screen "Inert Gas Conditioning Plant" 1280x800, template "Template_lite"
   on GenerateScreen: "TitleUpdater"()
   GraphicView "Graphic view_20" at 359,634 size 43x62; Picture "Graphic_72"
   GraphicView "Graphic view_52" at 746,80 size 58x108; Picture "Graphic_72"
   GraphicView "Graphic view_63" at 991,218 size 58x108; Picture "Graphic_72"
   GraphicView "Graphic view_64" at 1096,218 size 58x108; Picture "Graphic_72"
   TextField "Text field_64" at 497,462 size 54x22; Text '- OK -'
      Visibility <- "10_DI_DATA_LS_303_LO"
   GraphicView "Graphic view_76" at 53,433 size 168x182; Picture "Graphic_251"
   GraphicView "Graphic view_102" at 12,304 size 58x63; Picture "Graphic_162"
   GraphicView "Graphic view_13" at 724,163 size 182x22; Picture "Graphic_151"
   Group "Group" at 746,80 size 58x108; Picture "Graphic_72"
   GraphicIOField "Graphic I/O field_3" at 188,659 size 60x65; PictureList "Pump Ani"
      ProcessValue <- "10_DI_DATA_P_304_ENBLD"
   GraphicView "Graphic view_18" at 240,683 size 253x11; Picture "Graphic_156"
   GraphicView "Graphic view_89" at 303,257 size 10x13; Picture "Graphic_147"
   GraphicView "Graphic view_59" at 962,301 size 302x22; Picture "Graphic_151"
   GraphicView "Graphic view_5" at 827,163 size 102x22; Picture "Graphic_151"
   Group "Group_2" at 991,218 size 58x108; Picture "Graphic_72"
   TextField "Text field_45" at 989,239 size 60x22; Text 'Closed'
      Visibility <- "10_DI_DATA_CV407_CLSD"
   GraphicView "Graphic view_69" at 124,683 size 68x11; Picture "Graphic_156"
   GraphicView "Graphic view_85" at 235,296 size 33x35; Picture "Graphic_178"
   GraphicView "Graphic view_1" at 259,128 size 301x502; Picture "Graphic_150"
   GraphicView "Graphic view_6" at 870,257 size 18x22; Picture "Graphic_154"
   GraphicView "Graphic view_9" at 689,257 size 188x11; Picture "Graphic_156"
   GraphicView "Graphic view_11" at 424,625 size 12x91; Picture "Graphic_152"
   GraphicView "Graphic view_10" at 424,628 size 19x28; Picture "Graphic_157"
   GraphicView "Graphic view_12" at 440,636 size 106x11; Picture "Graphic_156"
   GraphicView "Graphic view_14" at 817,752 size 20x21; Picture "Graphic_159"
   GraphicView "Graphic view_16" at 635,761 size 188x13; Picture "Graphic_151"
   GraphicIOField "Graphic I/O field_1" at 573,615 size 60x65; PictureList "Pump Ani"
      ProcessValue <- "10_DI_DATA_P_303_ENBLD"
   GraphicView "Graphic view_19" at 471,636 size 106x11; Picture "Graphic_156"
   TextField "Text field_3" at 356,693 size 50x16; Text 'CV-358'
   Group "Group_1" at 359,634 size 43x62; Picture "Graphic_72"
   TextField "Text field_15" at 350,634 size 60x22; Text 'Closed'
      Visibility <- "10_DI_DATA_CV358_CLSD"
   TextField "Text field_16" at 90,573 size 90x22; Text 'PGC Running'
      Visibility <- "10_DI_DATA_E_400_RUN"
   GraphicView "Graphic view_21" at 486,674 size 17x18; Picture "Graphic_153"
   GraphicView "Graphic view_22" at 494,642 size 10x41; Picture "Graphic_152"
   GraphicView "Graphic view_23" at 490,637 size 17x15; Picture "Graphic_161"
   GraphicView "Graphic view_24" at 630,636 size 87x11; Picture "Graphic_156"
   GraphicView "Graphic view_30" at 421,704 size 39x47; Picture "Graphic_162"
   GraphicView "Graphic view_26" at 424,662 size 12x54; Picture "Graphic_152"
   TextField "Text field_1" at 460,713 size 60x22; Text 'Closed'
      Visibility <- "10_DI_DATA_CV341_CLSD"
   TextField "Text field_2" at 460,713 size 60x22; Text 'Opened'
      Visibility <- "10_DI_DATA_CV341_OPN"
   GraphicView "Graphic view_33" at 668,469 size 24x18; Picture "Graphic_155"
   GraphicView "Graphic view_34" at 668,508 size 24x18; Picture "Graphic_166"
   GraphicView "Graphic view_35" at 679,517 size 62x11; Picture "Graphic_156"
   GraphicView "Graphic view_36" at 668,486 size 12x30; Picture "Graphic_152"
   GraphicView "Graphic view_37" at 687,468 size 62x11; Picture "Graphic_156"
   GraphicView "Graphic view_38" at 741,468 size 106x11; Picture "Graphic_156"
   GraphicView "Graphic view_39" at 487,257 size 103x11; Picture "Graphic_156"
   GraphicView "Graphic view_40" at 422,102 size 140x11; Picture "Graphic_156"
   GraphicView "Graphic view_41" at 302,103 size 24x18; Picture "Graphic_155"
   GraphicView "Graphic view_43" at 558,103 size 19x18; Picture "Graphic_154"
   GraphicView "Graphic view_44" at 302,118 size 12x75; Picture "Graphic_152"
   GraphicView "Graphic view_45" at 302,183 size 12x75; Picture "Graphic_152"
   GraphicView "Graphic view_46" at 871,460 size 17x18; Picture "Graphic_153"
   GraphicView "Graphic view_47" at 879,426 size 10x41; Picture "Graphic_152"
   GraphicView "Graphic view_48" at 771,468 size 106x11; Picture "Graphic_156"
   GraphicView "Graphic view_49" at 879,358 size 10x91; Picture "Graphic_152"
   GraphicView "Graphic view_51" at 879,272 size 10x91; Picture "Graphic_152"
   GraphicView "Graphic view_53" at 574,257 size 126x11; Picture "Graphic_156"
   GraphicView "Graphic view_57" at 319,102 size 140x11; Picture "Graphic_156"
   TextField "Text field_4" at 434,743 size 50x16; Text 'CV-341'
   GraphicView "Graphic view_58" at 1062,188 size 19x119; Picture "Graphic_147"
   GraphicView "Graphic view_60" at 1058,159 size 58x63; Picture "Graphic_162"
   TextField "Text field_6" at 995,322 size 50x16; Text 'CV-407'
   GraphicView "Graphic view_61" at 561,250 size 23x16; Picture "Graphic_168"
   GraphicView "Graphic view_62" at 567,179 size 10x77; Picture "Graphic_152"
   TextField "Text field_8" at 1103,322 size 50x16; Text 'CV-411'
   Group "Group_3" at 1096,218 size 58x108; Picture "Graphic_72"
   GraphicView "Graphic view_65" at 1062,151 size 19x23; Picture "Graphic_147"
   TextField "Text field_9" at 1097,239 size 60x22; Text 'Closed'
      Visibility <- "10_DI_DATA_CV411_CLSD"
   TextField "Text field_10" at 1097,239 size 60x22; Text 'Opened'
      Visibility <- "10_DI_DATA_CV411_OPN"
   TextField "Text field_13" at 1115,180 size 60x22; Text 'Opened'
      Visibility <- "10_DI_DATA_CV409_OPN"
   TextField "Text field_17" at 582,680 size 42x16; Text 'P-303'
   TextField "Text field_5" at 1082,214 size 50x16; Text 'CV-409'
   GraphicView "Graphic view_66" at 508,761 size 188x13; Picture "Graphic_151"
   GraphicView "Graphic view_67" at 375,761 size 188x13; Picture "Graphic_151"
   GraphicView "Graphic view_31" at 424,748 size 12x38; Picture "Graphic_152"
   GraphicView "Graphic view_68" at 118,761 size 285x13; Picture "Graphic_151"
   GraphicView "Graphic view_70" at 826,617 size 12x146; Picture "Graphic_147"
   GraphicView "Graphic view_71" at 818,611 size 19x21; Picture "Graphic_169"
   GraphicView "Graphic view_73" at 14,359 size 19x222; Picture "Graphic_147"
   GraphicView "Graphic view_75" at 696,479 size 76x194; Picture "Graphic_173"
   GraphicView "Graphic view_72" at 760,610 size 68x13; Picture "Graphic_151"
   GraphicView "Graphic view_32" at 847,514 size 19x20; Picture "Graphic_169"
   GraphicView "Graphic view_77" at 759,513 size 97x13; Picture "Graphic_151"
   GraphicView "Graphic view_28" at 855,527 size 12x146; Picture "Graphic_147"
   GraphicView "Graphic view_79" at 855,649 size 12x130; Picture "Graphic_147"
   TextField "Text field_24" at 610,79 size 50x16; Text 'CV-405'
   TextField "Text field_27" at 820,266 size 48x16; Text 'FS-350'
   GraphicView "Graphic view_15" at 834,232 size 20x26; Picture "Graphic_79"
   TextField "Text field_40" at 813,209 size 70x22; Text 'No Flow'
      Visibility <- "10_DI_DATA_FS_350_FLW_OK"
   TextField "Text field_41" at 813,209 size 70x22; Text '- Flow -'
      Visibility <- "10_DI_DATA_FS_350_FLW_OK"
   GraphicView "Graphic view_8" at 558,596 size 10x11; Picture "Graphic_159"
   GraphicView "Graphic view_17" at 563,440 size 5x162; Picture "Graphic_147"
   GraphicView "Graphic view_25" at 558,275 size 10x11; Picture "Graphic_169"
   GraphicView "Graphic view_27" at 563,280 size 5x177; Picture "Graphic_147"
   GraphicView "Graphic view_29" at 486,602 size 78x5; Picture "Graphic_151"
   GraphicView "Graphic view_80" at 488,275 size 76x5; Picture "Graphic_151"
   IOField "I/O field_2" at 524,401 size 82x35; FormatPattern 999.9; Unit  %
      ProcessValue <- "12_AI_Data_LIT_304_SCALED"
   TextField "Text field_29" at 669,184 size 56x16; Text 'PIT-416'
   GraphicView "Graphic view_81" at 687,140 size 20x26; Picture "Graphic_36"
   TextField "Text field_25" at 752,442 size 56x16; Text 'TIT-408'
   TextField "Text field_30" at 512,199 size 56x16; Text 'TIT-406'
   GraphicView "Graphic view_82" at 530,137 size 20x26; Picture "Graphic_36"
   TextField "Text field_26" at 824,348 size 56x16; Text 'PIT-353'
   GraphicView "Graphic view_84" at 15,559 size 33x36; Picture "Graphic_177"
   TextField "Text field_7" at 750,184 size 50x16; Text 'CV-406'
   Bar "Bar_1" at 377,282 size 109x327; Unit  %; MinimumValue 0; MaximumValue 100
      ProcessValue <- "12_AI_Data_LIT_304_SCALED"
   TextField "Text field_48" at 16,624 size 112x20; Text 'PG Compressor'
      Appearance <- "10_DI_DATA_E_400_NOK"
   TextField "Text field_34" at 615,534 size 79x34; Text 'Heat Exchanger'
   TextField "Text field_35" at 551,697 size 100x34; Text 'Recirculation Pump'
   TextField "Text field_36" at 402,782 size 61x18; Text 'To Bilge'
   TextField "Text field_37" at 814,782 size 100x18; Text 'To Overboard'
   Group "Group_5" at 396,264 size 74x42
   GraphicView "Graphic view_3" at 429,258 size 15x16; Picture "Graphic_178"
   GraphicView "Graphic view_88" at 434,257 size 55x11; Picture "Graphic_151"
   TextField "Text field_38" at 571,440 size 55x16; Text 'LIT-304'
   TextField "Text field_39" at 269,693 size 56x16; Text 'PIT-358'
   GraphicView "Graphic view_90" at 287,658 size 20x26; Picture "Graphic_36"
   TextField "Text field_28" at 704,774 size 56x16; Text 'PIT-348'
   GraphicView "Graphic view_83" at 722,736 size 20x26; Picture "Graphic_36"
   TextField "Text field_31" at 778,623 size 48x16; Text 'FS-332'
   GraphicView "Graphic view_91" at 801,585 size 20x26; Picture "Graphic_79"
   TextField "Text field_32" at 779,562 size 70x22; Text 'No Flow'
      Visibility <- "10_DI_DATA_FS_332 FLW_OK"
   TextField "Text field_42" at 779,562 size 70x22; Text '- Flow -'
      Visibility <- "10_DI_DATA_FS_332 FLW_OK"
   TextField "Text field_43" at 197,724 size 42x16; Text 'P-304'
   TextField "Text field_44" at 169,740 size 106x20; Text 'Booster Pump'
   GraphicView "Graphic view_2" at 553,163 size 182x22; Picture "Graphic_151"
   TextField "Text field_11" at 989,239 size 60x22; Text 'Opened'
      Visibility <- "10_DI_DATA_CV407_OPN"
   GraphicView "Graphic view_7" at 251,453 size 24x21; Picture "Graphic_107"
   TextField "Text field_46" at 225,501 size 86x16; Text 'E-400-PT002'
   TextField "Text field_47" at 132,408 size 86x16; Text 'E-400-TT002'
   GraphicView "Graphic view_87" at 234,321 size 19x128; Picture "Graphic_147"
   GraphicView "Graphic view_86" at 220,442 size 33x36; Picture "Graphic_159"
   IOField "I/O field_10" at 683,53 size 57x22; FormatPattern 999
      ProcessValue <- "12_AI_Data_CV_405_SCALED"
   IOField "I/O field_11" at 226,482 size 68x18; FormatPattern 999.9; Unit  Bar
      ProcessValue <- "12_AI_Data_E_400_PT002_SCALED"
   IOField "I/O field_13" at 663,119 size 68x18; FormatPattern 99.99; Unit  Bar
      ProcessValue <- "12_AI_Data_PIT_416_SCALED"
   IOField "I/O field_14" at 787,330 size 68x18; FormatPattern 99.99; Unit  Bar
      ProcessValue <- "12_AI_Data_PIT_353_SCALED"
   IOField "I/O field_15" at 704,426 size 68x18; FormatPattern 99.99; Unit  °C
      ProcessValue <- "12_AI_Data_TIT_408_SCALED"
   IOField "I/O field_16" at 698,717 size 68x18; FormatPattern 99.99; Unit  Bar
      ProcessValue <- "12_AI_Data_PIT_348_SCALED"
   IOField "I/O field_7" at 263,638 size 68x18; FormatPattern 99.99; Unit  Bar
      ProcessValue <- "12_AI_Data_PIT_358_SCALED"
   TextField "Text field_57" at 1021,112 size 90x32; Text 'Vent To Atmosphere'
   TextField "Text field_58" at 608,3 size 150x18; Text 'Vent To Atmosphere'
   IOField "I/O field_1" at 143,392 size 68x18; FormatPattern 999.9; Unit  °C
      ProcessValue <- "12_AI_Data_E_400_TE002_SCALED"
   GraphicView "Graphic view_93" at 491,492 size 24x21; Picture "Graphic_107"
   TextField "Text field_63" at 515,491 size 48x16; Text 'LS-303'
   TextField "Text field_66" at 497,462 size 54x22; Text 'Low Low'
      Visibility <- "10_DI_DATA_LS_303_LO"
   TextField "Text field_90" at 497,462 size 54x22; Text '-LOW-'
      Visibility <- "10_DI_DATA_LS_303_LO"
   GraphicView "Graphic view_94" at 99,304 size 58x63; Picture "Graphic_162"
   TextField "Text field_70" at 125,264 size 60x22; Text 'Opened'
      Visibility <- "10_DI_DATA_CV441_OPN"
   TextField "Text field_71" at 126,288 size 50x16; Text 'CV-441'
   GraphicView "Graphic view_95" at 103,278 size 19x41; Picture "Graphic_147"
   TextField "Text field_72" at 93,222 size 65x32; Text 'Ambient Air Inlet'
   GraphicView "Graphic view_96" at 86,364 size 36x39; Picture "Graphic_159"
   GraphicView "Graphic view_97" at 28,382 size 70x22; Picture "Graphic_151"
   TextField "Text field_69" at 125,264 size 60x22; Text 'Closed'
      Visibility <- "10_DI_DATA_CV441_CLSD"
   TextField "Text field_12" at 1115,180 size 60x22; Text 'Closed'
      Visibility <- "10_DI_DATA_CV409_CLSD"
   GraphicView "Graphic view_98" at 0,278 size 33x35; Picture "Graphic_169"
   GraphicView "Graphic view_99" at 856,330 size 23x20; Picture "Graphic_255"
   GraphicView "Graphic view_100" at 728,443 size 20x26; Picture "Graphic_36"
   TextField "Text field_33" at 744,96 size 60x22; Text 'Closed'
      Visibility <- "10_DI_DATA_CV406_CLSD"
   TextField "Text field_14" at 744,96 size 60x22; Text 'Opened'
      Visibility <- "10_DI_DATA_CV406_OPN"
   TextField "Text field_18" at 950,356 size 149x23; Text 'Hazardous Area'
   GraphicView "Graphic view_4" at 1204,277 size 20x26; Picture "Graphic_36"
   IOField "I/O field_3" at 1180,257 size 68x18; FormatPattern 99.99; Unit  Bar
      ProcessValue <- "20_TANKS_IP_DATA_RIO_06_FIRST_TANK_DECK_IG_PRESS"
   TextField "Text field_20" at 1186,322 size 56x16; Text 'PIT-415'
   GraphicView "Graphic view_50" at 100,253 size 26x26; Picture "Graphic_261"
   GraphicView "Graphic view_74" at 549,146 size 18x54; Picture "Graphic_281"
   GraphicView "Graphic view_78" at 256,278 size 17x59; Picture "Graphic_281"
   GraphicView "Graphic view_101" at 213,397 size 23x20; Picture "Graphic_255"
   TextField "Text field_56" at 1229,342 size 44x32; Text 'To BWTS'
   TextField "Text field_60" at 661,356 size 94x23; Text 'Safe Area'
   IOField "I/O field_4" at 683,37 size 57x22; FormatPattern 999
      ProcessValue <- "16_AQ_Data_CV405_CNTRL"
   TextField "Text field_106" at 752,38 size 59x18; Text 'OPENED'
   GraphicView "Graphic view_103" at 14,298 size 19x22; Picture "Graphic_147"
   TextField "Text field_73" at 34,288 size 50x16; Text 'CV-401'
   TextField "Text field_74" at 30,264 size 60x22; Text 'Opened'
      Visibility <- "10_DI_Data_CV401_OPN"
   TextField "Text field_75" at 30,264 size 60x22; Text 'Closed'
      Visibility <- "10_DI_Data_CV401_CLSD"
   Button "HmiScreenItemData_13" at 4,669 size 121x40; TextOn 'IGG Plant'; TextOff 'Fresh Water System'; Authorization "Operate"
      on Release: ActivateScreen("Fresh Water System", 0)
      Appearance <- "10 DI_DATA_P305_ENBLD"
   Button "HmiScreenItemData_11" at 3,745 size 122x41; TextOn 'IGG Plant'; TextOff 'Cooling System'; Authorization "Operate"
      on Release: ActivateScreen("Cooling System", 0)
   TextField "Text field_22" at 90,573 size 90x22; Text 'PGC Loaded'
      Visibility <- "10_DI_DATA_E_400_RUN"
   Button "HmiScreenItemData_12" at 46,424 size 177x198; TextOn 'IGG Plant'; TextOff 'Text'; Authorization "Operate"
      on Release: ActivateScreen("PGC System", 0)
   TextField "Text field_23" at 350,634 size 60x22; Text 'Opened'
      Visibility <- "10_DI_DATA_CV358_OPN"
   GraphicView "Graphic view_54" at 588,60 size 19x108; Picture "Graphic_147"
   GraphicView "Graphic view_55" at 586,28 size 95x54; Picture "Graphic_167"
   GraphicView "Graphic view_56" at 588,8 size 19x33; Picture "Graphic_147"
   IOField "I/O field_12" at 506,119 size 68x18; FormatPattern 99.99; Unit  °C
      ProcessValue <- "12_AI_Data_TIT_406_SCALED"
   GraphicView "Graphic view_42" at 567,116 size 10x51; Picture "Graphic_152"
   TextField "Text field_76" at 618,40 size 30x22; Text 'A'
      Visibility <- "19_AUTO_CMNDS_Data_CV405_PID_MDLTG"
   GraphicView "Logo" at 1,1 size 219x60; Picture "Logo of IGG HMI"
   Button "HmiScreenItemData_1" at 1,50 size 150x43; TextOn 'Back'; TextOff 'Main Index'
      on Release: ActivateScreen("02 Main Index", 0)
   GraphicView "Graphic view_92" at 925,164 size 33x36; Picture "Graphic_169"
   Button "HmiScreenItemData_2" at 1128,64 size 150x43; TextOn 'Back'; TextOff 'GCU Setup'; Authorization "Operate"
      on Release: ActivateScreen("Inert Gas Conditioning Setup", 0)
   DateTimeField "HmiScreenItemData_17" at 1175,0 size 105x30
   DateTimeField "HmiScreenItemData" at 1175,30 size 105x30
   GraphicView "Graphic view_106" at 939,194 size 19x100; Picture "Graphic_147"
   GraphicView "Graphic view_104" at 940,285 size 33x37; Picture "Graphic_177"
   Button "HmiScreenItemData_9" at 930,410 size 340x30; TextOn 'Back'; TextOff 'GCU CONTROL'
      Visibility <- "150_GCU_LCL_CNTRL_DB_LCL_CNTRL_ACTV"
   Line "Line_2" at 1246,550 size 0x80
      Visibility <- "150_GCU_LCL_CNTRL_DB_LCL_CNTRL_ACTV"
   Line "Line_3" at 1080,630 size 166x0
      Visibility <- "150_GCU_LCL_CNTRL_DB_LCL_CNTRL_ACTV"
   Button "HmiScreenItemData_4" at 930,610 size 150x40; TextOn 'Back'; TextOff 'Stop'; Authorization "Commissioning"
      on Press: function_b14e0dd5("150_GCU_LCL_CNTRL_DB_STOP", 0)
      Visibility <- "150_GCU_LCL_CNTRL_DB_LCL_CNTRL_ACTV"
   Line "Line_7" at 1080,530 size 145x0
      Visibility <- "150_GCU_LCL_CNTRL_DB_LCL_CNTRL_ACTV"
   Circle "Circle_20" at 1225,510 size 40x40
      Visibility <- "150_GCU_LCL_CNTRL_DB_LCL_CNTRL_ACTV"
      Appearance <- "150_GCU_LCL_CNTRL_DB_RUN_WITH_AIR"
   Button "HmiScreenItemData_3" at 930,510 size 150x40; TextOn 'Back'; TextOff 'Start With Air'; Authorization "Commissioning"
      on Press: function_b14e0dd5("150_GCU_LCL_CNTRL_DB_STRT_AIR", 0)
      Visibility <- "150_GCU_LCL_CNTRL_DB_LCL_CNTRL_ACTV"
   Button "HmiScreenItemData_5" at 930,450 size 340x40; TextOn 'Back'; TextOff 'Start'; TextList "GCU_LCL"; Authorization "Commissioning"
      on Press: InvertBit("150_GCU_LCL_CNTRL_DB_LCL_CNTRL_ACTV")
      Visibility <- "150_GCU_LCL_CNTRL_DB_LCL_CNTRL_ACTV"
      ProcessValue <- "150_GCU_LCL_CNTRL_DB_LCL_CNTRL_ACTV"
   Button "HmiScreenItemData_6" at 930,560 size 150x40; TextOn 'Back'; TextOff 'Start With IG'; Authorization "Commissioning"
      on Press: function_b14e0dd5("150_GCU_LCL_CNTRL_DB_STRT_IG", 0)
      Visibility <- "150_GCU_LCL_CNTRL_DB_LCL_CNTRL_ACTV"
   Line "Line_6" at 1080,580 size 145x0
      Visibility <- "150_GCU_LCL_CNTRL_DB_LCL_CNTRL_ACTV"
   Circle "Circle_1" at 1225,560 size 40x40
      Visibility <- "150_GCU_LCL_CNTRL_DB_LCL_CNTRL_ACTV"
      Appearance <- "150_GCU_LCL_CNTRL_DB_RUN_WITH_IG"
   Button "HmiScreenItemData_7" at 930,660 size 240x40; TextOn 'Back'; TextOff 'Start With Air'; TextList "GTT_OPS"; Authorization "Commissioning"
      on Press: InvertBit("150_GCU_LCL_CNTRL_DB_OPN_ACTV_GTT_VLVS")
      Visibility <- "150_GCU_LCL_CNTRL_DB_LCL_CNTRL_ACTV"
      ProcessValue <- "150_GCU_LCL_CNTRL_DB_OPN_ACTV_GTT_VLVS"
   Circle "Circle_2" at 1225,660 size 40x40
      Visibility <- "150_GCU_LCL_CNTRL_DB_LCL_CNTRL_ACTV"
      Appearance <- "150_GCU_LCL_CNTRL_DB_OPN_ACTV_GTT_VLVS"
   Line "Line_14" at 1170,680 size 55x0
      Visibility <- "150_GCU_LCL_CNTRL_DB_LCL_CNTRL_ACTV"
   Group "Group_4" at 187,631 size 60x25
   Group "Group_6" at 573,588 size 60x25
   IOField "I/O field_34" at 664,96 size 66x23; FormatPattern 99.9; Unit  Bar
      ProcessValue <- "19_AUTO_CMNDS_Data_PIT416_CMND_Target"
      Appearance <- "19_AUTO_CMNDS_Data_PIT402_Target"
   Group "Group_7" at 214,1 size 373x50
   GraphicView "Graphic view_105" at 1184,288 size 96x48; Picture "Graphic_235"
   Button "HmiScreenItemData_10" at 1178,277 size 102x71; TextOn 'Back'; TextOff 'Text'
      on Press: ActivateScreen("Balast Water Treatment Plant", 0)
   GraphicView "Graphic view_108" at 2,208 size 95x48; Picture "Left Arow"
   Button "HmiScreenItemData_14" at 1,195 size 106x107; TextOn 'Back'; TextOff 'Text'
      on Press: ActivateScreen("Inert Gas Generator Plant", 0)
   Button "HmiScreenItemData_15" at 1,133 size 158x52; TextOn 'INERT GAS TRANSFER'; TextOff 'Inert Gas Transfer'; TextList "IG Transfer"; Authorization "Operate"
      on Release: ActivateScreen("IG Transfer Mode", 0)
      ProcessValue <- "80_From_HMI_BWT_BYPASS"
   IOField "I/O field_37" at 1070,718 size 79x29; Authorization "Commissioning"; FormatPattern 999; Unit  step
      ProcessValue <- "2110_BTCS_CNTRL_DB_BTCS_STEP"
   Button "HmiScreenItemData_16" at 930,718 size 137x29; TextOn 'Back'; TextOff 'BWTS Step'
   Button "HmiScreenItemData_51" at 930,753 size 137x29; TextOn 'Back'; TextOff 'BWTS State'
   IOField "I/O field_38" at 1070,753 size 79x29; Authorization "Commissioning"; FormatPattern 9; Unit  state
      ProcessValue <- "2110_BTCS_CNTRL_DB_BTCS_STATE"
   Group "Group_9" at 591,11 size 604x305
   Group "Group_12" at 260,515 size 606x260
   Group "Group_13" at 179,634 size 324x58
   GraphicView "Graphic view_107" at 563,347 size 57x58; Picture "Graphic_302"
      Visibility <- "10_DI_DATA_EPB_8S1"
   Group "Group_10" at 389,152 size 96x105
   Group "Group_11" at 239,299 size 243x195
   Group "Group_8" at 384,257 size 504x388
   Button "Button_1" at 655,120 size 84x92; TextOff 'Text'
      on Press: function_efd93a16("PGC Setpoint Protection", 400, 200, -1, -1, 1)
   Button "Button_4" at 578,3 size 84x99; TextOff 'Text'
      on Press: function_efd93a16("CV 405 Grafics", 300, 100, -1, -1, 1)
   Button "HmiScreenItemData_18" at 236,593 size 83x29; TextOn 'Back'; TextOff 'Temp-Trends'
      on Click: function_efd93a16("PGC Temperature Trends", 200, 100, -1, -1, 1)
   Group "Group_14" at 914,406 size 366x378
   Button "Button_3" at 187,631 size 60x25; TextOn 'Alarm'; TextOff 'OK'
      Appearance <- "10_DI_DATA_P_304_OK"
   TextField "Text field_19" at 187,631 size 60x25; Text 'Enabled'
      Visibility <- "14_DQ_DATA_P_304"
      Appearance <- "14_DQ_DATA_P_304"
   Button "Button_2" at 573,588 size 60x25; TextOn 'Alarm'; TextOff 'OK'
      Appearance <- "10_DI_DATA_P_303_OK"
   TextField "Text field_49" at 573,588 size 60x25; Text 'Enabled'
      Visibility <- "14_DQ_DATA_P_303"
      Appearance <- "14_DQ_DATA_P_303"
   Button "HmiScreenItemData_8" at 228,5 size 355x40; TextOn 'Back'; TextOff 'Text'
   TextField "Screen title" at 214,1 size 373x50; Text 'Screen title'
   Circle "Circle_73" at 594,11 size 10x10
      VerticalMovement <- "E-400 Animation_DB_Animation"
      Visibility <- "10_DI_DATA_E_400_RUN"
   Circle "Circle_45" at 592,89 size 10x10
      VerticalMovement <- "E-400 Animation_DB_Animation"
      Visibility <- "10_DI_DATA_E_400_RUN"
   Circle "Circle_84" at 591,169 size 10x10
      HorizontalMovement <- "E-400 Animation_DB_Animation"
      Visibility <- "10_DI_DATA_E_400_RUN"
   Circle "Circle_26" at 706,169 size 10x10
      HorizontalMovement <- "E-400 Animation_DB_Animation"
      Visibility <- "10_DI_DATA_CV406_CLSD"
   Circle "Circle_27" at 748,169 size 10x10
      HorizontalMovement <- "E-400 Animation_DB_Animation"
      Visibility <- "10_DI_DATA_CV406_CLSD"
   Circle "Circle_28" at 811,169 size 10x10
      HorizontalMovement <- "E-400 Animation_DB_Animation"
      Visibility <- "10_DI_DATA_CV407_CLSD"
   Circle "Circle_29" at 876,169 size 10x10
      HorizontalMovement <- "E-400 Animation_DB_Animation"
      Visibility <- "10_DI_DATA_CV407_CLSD"
   Circle "Circle_72" at 882,168 size 10x10
      HorizontalMovement <- "E-400 Animation_DB_Animation"
      Visibility <- "10_DI_DATA_CV407_CLSD"
   Circle "Circle_30" at 929,168 size 10x10
      HorizontalMovement <- "E-400 Animation_DB_Animation"
      Visibility <- "10_DI_DATA_CV407_CLSD"
   Circle "Circle_71" at 940,168 size 10x10
      HorizontalMovement <- "E-400 Animation_DB_Animation"
      Visibility <- "10_DI_DATA_CV407_CLSD"
   Circle "Circle_31" at 944,304 size 10x10
      VerticalMovement <- "E-400 Animation_DB_Animation"
      Visibility <- "10_DI_DATA_CV407_CLSD"
   Circle "Circle_42" at 995,305 size 10x10
      HorizontalMovement <- "E-400 Animation_DB_Animation"
      Visibility <- "10_DI_DATA_CV407_CLSD"
   Circle "Circle_44" at 1066,143 size 10x10
      VerticalMovement <- "E-400 Animation_DB_Animation"
      Visibility <- "10_DI_DATA_CV409_CLSD"
   Circle "Circle_43" at 1066,224 size 10x10
      VerticalMovement <- "E-400 Animation_DB_Animation"
      Visibility <- "10_DI_DATA_CV409_CLSD"
   Circle "Circle_32" at 1098,306 size 10x10
      HorizontalMovement <- "E-400 Animation_DB_Animation"
      Visibility <- "10_DI_DATA_CV411_CLSD"
   Circle "Circle_82" at 1185,305 size 10x10
      HorizontalMovement <- "E-400 Animation_DB_Animation"
      Visibility <- "10_DI_DATA_CV411_CLSD"
   Circle "Circle_67" at 260,764 size 8x8
      Visibility <- "10_DI_DATA_FS_332 FLW_OK"
      HorizontalMovement <- "FS332 Animation_IDB_Animation"
   Circle "Circle_68" at 411,763 size 8x8
      Visibility <- "10_DI_DATA_FS_332 FLW_OK"
      HorizontalMovement <- "FS332 Animation_IDB_Animation"
   Circle "Circle_69" at 573,764 size 8x8
      Visibility <- "10_DI_DATA_FS_332 FLW_OK"
      HorizontalMovement <- "FS332 Animation_IDB_Animation"
   Circle "Circle_70" at 712,763 size 8x8
      Visibility <- "10_DI_DATA_FS_332 FLW_OK"
      HorizontalMovement <- "FS332 Animation_IDB_Animation"
   Circle "Circle_74" at 813,763 size 8x8
      Visibility <- "10_DI_DATA_FS_332 FLW_OK"
      HorizontalMovement <- "FS332 Animation_IDB_Animation"
   Circle "Circle_75" at 828,691 size 8x8
      Visibility <- "10_DI_DATA_FS_332 FLW_OK"
      VerticalMovement <- "FS332 Animation_IDB_Animation"
   Circle "Circle_76" at 828,633 size 8x8
      Visibility <- "10_DI_DATA_FS_332 FLW_OK"
      VerticalMovement <- "FS332 Animation_IDB_Animation"
   Circle "Circle_77" at 763,613 size 8x8
      Visibility <- "10_DI_DATA_FS_332 FLW_OK"
      HorizontalMovement <- "FS332 Animation_IDB_Animation"
   Circle "Circle_78" at 845,515 size 10x10
      Visibility <- "10_DI_DATA_FS_332 FLW_OK"
      HorizontalMovement <- "FS332 Animation_IDB_Animation"
   Circle "Circle_79" at 856,642 size 10x10
      Visibility <- "10_DI_DATA_FS_332 FLW_OK"
      VerticalMovement <- "FS332 Animation_IDB_Animation"
   Circle "Circle_80" at 856,765 size 10x10
      Visibility <- "10_DI_DATA_FS_332 FLW_OK"
      VerticalMovement <- "FS332 Animation_IDB_Animation"
   Circle "Circle_55" at 179,684 size 7x7
      HorizontalMovement <- "P304 Animation_IDB_Animation"
      Visibility <- "10_DI_DATA_CV358_OPN"
   Circle "Circle_83" at 318,685 size 7x7
      DiagonalMovement <- "P304 Animation_IDB_Animation"
      Visibility <- "10_DI_DATA_CV358_OPN"
   Circle "Circle_81" at 416,684 size 7x7
      DiagonalMovement <- "P304 Animation_IDB_Animation"
      Visibility <- "10_DI_DATA_CV358_OPN"
   Circle "Circle_56" at 485,684 size 7x7
      DiagonalMovement <- "P304 Animation_IDB_Animation"
      Visibility <- "10_DI_DATA_CV358_OPN"
   Circle "Circle_85" at 496,641 size 7x7
      DiagonalMovement <- "P304 Animation_IDB_Animation"
      Visibility <- "10_DI_DATA_CV358_OPN"
   Circle "Circle_86" at 426,634 size 7x7
      DiagonalMovement <- "P304 Animation_IDB_Animation"
      Visibility <- "10_DI_DATA_CV358_OPN"
   Circle "Circle_38" at 389,247 size 9x9
      DiagonalMovement <- "E-400 Animation_DB_Animation"
      Visibility <- "10_DI_DATA_E_400_RUN"
   Circle "Circle_57" at 402,247 size 10x10
      DiagonalMovement <- "E-400 Animation_DB_Animation"
      Visibility <- "10_DI_DATA_E_400_RUN"
   Circle "Circle_40" at 417,247 size 10x10
      DiagonalMovement <- "E-400 Animation_DB_Animation"
      Visibility <- "10_DI_DATA_E_400_RUN"
   Circle "Circle_58" at 433,247 size 10x10
      DiagonalMovement <- "E-400 Animation_DB_Animation"
      Visibility <- "10_DI_DATA_E_400_RUN"
   Circle "Circle_60" at 475,162 size 10x10
      DiagonalMovement <- "E-400 Animation_DB_Animation"
      Visibility <- "10_DI_DATA_E_400_RUN"
   Circle "Circle_41" at 474,180 size 10x10
      DiagonalMovement <- "E-400 Animation_DB_Animation"
      Visibility <- "10_DI_DATA_E_400_RUN"
   Circle "Circle_39" at 475,172 size 9x9
      DiagonalMovement <- "E-400 Animation_DB_Animation"
      Visibility <- "10_DI_DATA_E_400_RUN"
   Circle "Circle_59" at 475,152 size 10x10
      DiagonalMovement <- "E-400 Animation_DB_Animation"
      Visibility <- "10_DI_DATA_E_400_RUN"
   Circle "Circle_87" at 448,247 size 10x10
      DiagonalMovement <- "E-400 Animation_DB_Animation"
      Visibility <- "10_DI_DATA_E_400_RUN"
   Circle "Circle_88" at 462,247 size 10x10
      DiagonalMovement <- "E-400 Animation_DB_Animation"
      Visibility <- "10_DI_DATA_E_400_RUN"
   Circle "Circle_89" at 474,190 size 10x10
      DiagonalMovement <- "E-400 Animation_DB_Animation"
      Visibility <- "10_DI_DATA_E_400_RUN"
   Circle "Circle_90" at 474,199 size 10x10
      DiagonalMovement <- "E-400 Animation_DB_Animation"
      Visibility <- "10_DI_DATA_E_400_RUN"
   Circle "Circle_33" at 239,444 size 10x10
      DiagonalMovement <- "E-400 Animation_DB_Animation"
      Visibility <- "10_DI_DATA_E_400_RUN"
   Circle "Circle_34" at 240,306 size 11x11
      Visibility <- "10_DI_DATA_E_400_RUN"
      VerticalMovement <- "E-400 Animation_DB_Animation"
   Circle "Circle_35" at 307,299 size 12x12
      Visibility <- "10_DI_DATA_E_400_RUN"
      HorizontalMovement <- "E-400 Animation_DB_Animation"
   Circle "Circle_36" at 308,423 size 12x12
      DiagonalMovement <- "E-400 Animation_DB_Animation"
      Visibility <- "10_DI_DATA_E_400_RUN"
   Circle "Circle_37" at 357,481 size 13x13
      DiagonalMovement <- "E-400 Animation_DB_Animation"
      Visibility <- "10_DI_DATA_E_400_RUN"
   Circle "Circle_61" at 392,416 size 10x10
      DiagonalMovement <- "E-400 Animation_DB_Animation"
      Visibility <- "10_DI_DATA_E_400_RUN"
   Circle "Circle_63" at 408,416 size 10x10
      DiagonalMovement <- "E-400 Animation_DB_Animation"
      Visibility <- "10_DI_DATA_E_400_RUN"
   Circle "Circle_64" at 424,416 size 10x10
      DiagonalMovement <- "E-400 Animation_DB_Animation"
      Visibility <- "10_DI_DATA_E_400_RUN"
   Circle "Circle_65" at 456,416 size 10x10
      DiagonalMovement <- "E-400 Animation_DB_Animation"
      Visibility <- "10_DI_DATA_E_400_RUN"
   Circle "Circle_66" at 472,416 size 10x10
      DiagonalMovement <- "E-400 Animation_DB_Animation"
      Visibility <- "10_DI_DATA_E_400_RUN"
   Circle "Circle_62" at 440,416 size 10x10
      DiagonalMovement <- "E-400 Animation_DB_Animation"
      Visibility <- "10_DI_DATA_E_400_RUN"
   Circle "Circle_54" at 384,309 size 7x7
      DiagonalMovement <- "82_To_HMI_FS350 Animation"
      Visibility <- "10_DI_DATA_FS_350_FLW_OK"
   Circle "Circle_53" at 388,321 size 8x8
      DiagonalMovement <- "82_To_HMI_FS350 Animation"
      Visibility <- "10_DI_DATA_FS_350_FLW_OK"
   Circle "Circle_51" at 408,332 size 6x6
      DiagonalMovement <- "82_To_HMI_FS350 Animation"
      Visibility <- "10_DI_DATA_FS_350_FLW_OK"
   Circle "Circle_49" at 432,336 size 6x6
      DiagonalMovement <- "82_To_HMI_FS350 Animation"
      Visibility <- "10_DI_DATA_FS_350_FLW_OK"
   Circle "Circle_50" at 453,328 size 7x7
      DiagonalMovement <- "82_To_HMI_FS350 Animation"
      Visibility <- "10_DI_DATA_FS_350_FLW_OK"
   Circle "Circle_52" at 466,317 size 8x8
      DiagonalMovement <- "82_To_HMI_FS350 Animation"
      Visibility <- "10_DI_DATA_FS_350_FLW_OK"
   Circle "Circle_48" at 476,306 size 7x7
      DiagonalMovement <- "82_To_HMI_FS350 Animation"
      Visibility <- "10_DI_DATA_FS_350_FLW_OK"
   Circle "Circle_14" at 437,257 size 10x10
      DiagonalMovement <- "82_To_HMI_FS350 Animation"
      Visibility <- "10_DI_DATA_FS_350_FLW_OK"
   Circle "Circle_5" at 527,257 size 9x9
      DiagonalMovement <- "82_To_HMI_FS350 Animation"
      Visibility <- "10_DI_DATA_FS_350_FLW_OK"
   Circle "Circle_6" at 589,257 size 9x9
      DiagonalMovement <- "82_To_HMI_FS350 Animation"
      Visibility <- "10_DI_DATA_FS_350_FLW_OK"
   Circle "Circle_7" at 664,257 size 9x9
      DiagonalMovement <- "82_To_HMI_FS350 Animation"
      Visibility <- "10_DI_DATA_FS_350_FLW_OK"
   Circle "Circle_8" at 739,257 size 10x10
      DiagonalMovement <- "82_To_HMI_FS350 Animation"
      Visibility <- "10_DI_DATA_FS_350_FLW_OK"
   Circle "Circle_9" at 816,258 size 9x9
      DiagonalMovement <- "82_To_HMI_FS350 Animation"
      Visibility <- "10_DI_DATA_FS_350_FLW_OK"
   Circle "Circle_12" at 877,264 size 10x10
      Visibility <- "10_DI_DATA_FS_350_FLW_OK"
      VerticalMovement <- "82_To_HMI_FS350 Animation"
   Circle "Circle_13" at 878,359 size 10x10
      Visibility <- "10_DI_DATA_FS_350_FLW_OK"
      VerticalMovement <- "82_To_HMI_FS350 Animation"
   Circle "Circle_11" at 870,466 size 10x10
      DiagonalMovement <- "82_To_HMI_FS350 Animation"
      Visibility <- "10_DI_DATA_FS_350_FLW_OK"
   Circle "Circle_10" at 774,469 size 9x9
      DiagonalMovement <- "82_To_HMI_FS350 Animation"
      Visibility <- "10_DI_DATA_FS_350_FLW_OK"
   Circle "Circle_47" at 669,474 size 10x10
      Visibility <- "10_DI_DATA_FS_350_FLW_OK"
      VerticalMovement <- "82_To_HMI_FS350 Animation"
   Circle "Circle_46" at 667,509 size 10x10
      DiagonalMovement <- "82_To_HMI_FS350 Animation"
      Visibility <- "10_DI_DATA_FS_350_FLW_OK"
   Circle "Circle_15" at 475,635 size 10x10
      Visibility <- "10_DI_DATA_FS_350_FLW_OK"
      HorizontalMovement <- "82_To_HMI_FS350 Animation"
   Circle "Circle_16" at 518,635 size 10x10
      Visibility <- "10_DI_DATA_FS_350_FLW_OK"
      HorizontalMovement <- "82_To_HMI_FS350 Animation"
   Circle "Circle_17" at 562,635 size 10x10
      Visibility <- "10_DI_DATA_FS_350_FLW_OK"
      HorizontalMovement <- "82_To_HMI_FS350 Animation"
   Circle "Circle_18" at 661,635 size 9x9
      Visibility <- "10_DI_DATA_FS_350_FLW_OK"
      HorizontalMovement <- "82_To_HMI_FS350 Animation"
   Circle "Circle_19" at 684,635 size 9x9
      Visibility <- "10_DI_DATA_FS_350_FLW_OK"
      HorizontalMovement <- "82_To_HMI_FS350 Animation"
   Circle "Circle_21" at 403,292 size 6x6
      DiagonalMovement <- "82_To_HMI_FS350 Animation"
      Visibility <- "10_DI_DATA_FS_350_FLW_OK"
   Circle "Circle_22" at 410,301 size 6x6
      DiagonalMovement <- "82_To_HMI_FS350 Animation"
      Visibility <- "10_DI_DATA_FS_350_FLW_OK"
   Circle "Circle_25" at 418,306 size 6x6
      DiagonalMovement <- "82_To_HMI_FS350 Animation"
      Visibility <- "10_DI_DATA_FS_350_FLW_OK"
   Circle "Circle_3" at 429,307 size 7x7
      DiagonalMovement <- "82_To_HMI_FS350 Animation"
      Visibility <- "10_DI_DATA_FS_350_FLW_OK"
   Circle "Circle_4" at 445,307 size 5x5
      DiagonalMovement <- "82_To_HMI_FS350 Animation"
      Visibility <- "10_DI_DATA_FS_350_FLW_OK"
   Circle "Circle_23" at 453,302 size 5x5
      DiagonalMovement <- "82_To_HMI_FS350 Animation"
      Visibility <- "10_DI_DATA_FS_350_FLW_OK"
   Circle "Circle_24" at 460,295 size 6x6
      DiagonalMovement <- "82_To_HMI_FS350 Animation"
      Visibility <- "10_DI_DATA_FS_350_FLW_OK"
   TextField "Text field_50" at 969,420 size 254x154; Text 'Please Make Sure the Energy and Water Supply are Present and Sufficient'
      Visibility <- "Warn To Start GCU-Last"
   Button "Button_5" at 928,406 size 343x378; TextOff 'Text'
      Visibility <- "Warn To Start GCU-Last"
   TextField "Text field_21" at 919,606 size 359x94; Text 'Instalation Start Confirmation Required for Re-Ox Stage'
      Visibility <- "Warn To Start GCU-Last"
   Button "Button_6" at 1004,717 size 200x55; TextOff 'CONFIRM'; Authorization "Operate"
      on Press: function_b14e0dd5("80_From_HMI_GCU Start Confirmed", 0)
      Visibility <- "Warn To Start GCU-Last"
   TextField "Text field_51" at 914,433 size 366x124; Text 'Please Make Sure the Energy and Water Supply are Present and Sufficient'
      Visibility <- "Warn To Start GCU-Last"

screen "Balast Water Treatment Plant" 1280x800, template "Template"
   on GenerateScreen: "User_Change"(); "TitleUpdater"()
   Button "HmiScreenItemData_1" at 1,1 size 150x40; TextOn 'Back'; TextOff 'Main Index'
      on Release: ActivateScreen("02 Main Index", 0)
   TextField "Text field_63" at 383,107 size 72x30; Text 'Pre Dwell Time'
   Circle "Circle_29" at 1047,85 size 20x20
      Appearance <- "2102_TIME_CALCS_DB_POST_DWELL_TMR_DN"
   Button "HmiScreenItemData_9" at 10,60 size 158x27; TextOn 'Back'; TextOff 'BWTS Control'
   Button "HmiScreenItemData_4" at 14,150 size 75x47; TextOn 'Back'; TextOff 'Stop'; Authorization "Operate"
      on Release: function_efd93a16("BWTS Stop Confirm", 400, 200, -1, -1, 1)
      ObjectEnable <- "82_To_HMI_CRNT_MODE_GCU"
   Circle "Circle_20" at 137,105 size 29x29
      Appearance <- "82_To_HMI_IGG RUN Indication"
   Button "HmiScreenItemData_3" at 14,93 size 75x47; TextOn 'Back'; TextOff 'Start'; Authorization "Operate"
      on Release: function_efd93a16("BWTS Start Confirm", 400, 200, -1, -1, 1)
      ObjectEnable <- "82_To_HMI_CRNT_MODE_GCU"
   Button "HmiScreenItemData_2" at 1129,1 size 150x40; TextOn 'Back'; TextOff 'BWTS Setup'
      on Release: ActivateScreen("Balast Water Treatment Setup", 0)
   TextField "Text field_1" at 290,107 size 68x30; Text 'Tank Selected'
   TextField "Text field_2" at 841,107 size 61x30; Text 'BWTS Started'
   TextField "Text field_3" at 568,107 size 62x30; Text 'IGGS Started'
   TextField "Text field_4" at 659,107 size 60x30; Text 'GCU Started'
   TextField "Text field_5" at 748,107 size 61x30; Text 'PGC Started'
   TextField "Text field_6" at 908,107 size 102x30; Text 'Gas Transfer Started'
   Circle "Circle_10" at 956,89 size 14x14
      Appearance <- "2110_BTCS_CNTRL_DB_BTCS_STEP"
   TextField "Text field_7" at 995,107 size 125x30; Text 'Treatment Cycle Completed'
   TextField "Text field_21" at 306,401 size 54x20; Text 'Closed'
      Visibility <- "20_TANKS_IP_DATA_RIO_06_FIRST_TANK_GTT_ISOL_VALVE_CLSD"
   TextField "Text field_22" at 306,401 size 54x20; Text 'Opened'
      Visibility <- "20_TANKS_IP_DATA_RIO_06_FIRST_TANK_GTT_ISOL_VALVE_OPEN"
   GraphicView "Graphic view_10" at 283,396 size 22x31; Picture "Graphic_162"
   TextField "Text field_25" at 306,482 size 54x20; Text 'Closed'
      Visibility <- "20_TANKS_IP_DATA_RIO_06_SECOND_TANK_GTT_ISOL_VALVE_CLSD"
   TextField "Text field_26" at 306,482 size 54x20; Text 'Opened'
      Visibility <- "20_TANKS_IP_DATA_RIO_06_SECOND_TANK_GTT_ISOL_VALVE_OPEN"
   IOField "I/O field_2" at 309,560 size 72x20; FormatPattern 999; Unit Nm³/hr
      ProcessValue <- "20_TANKS_IP_DATA_RIO_06_SECOND_TANK_USD_FLOW"
   IOField "I/O field_4" at 309,599 size 72x20; FormatPattern 999; Unit Nm³/hr
      ProcessValue <- "20_TANKS_IP_DATA_RIO_06_SECOND_TANK_MBG_FLOW"
   TextField "Text field_27" at 263,602 size 29x14; Text 'MBG'
   TextField "Text field_28" at 285,545 size 33x15; Text 'USD'
   TextField "Text field_23" at 261,291 size 34x14; Text 'MBG'
   TextField "Text field_24" at 284,349 size 28x14; Text 'USD'
   Group "Group" at 1064,419 size 35x38; Picture "Graphic_72"
   TextField "Text field_19" at 1057,414 size 54x20; Text 'Closed'
      Visibility <- "20_TANKS_IP_DATA_RIO_01_FIRST_TANK_GTT_ISOL_VALVE_CLSD"
   TextField "Text field_20" at 1057,414 size 54x20; Text 'Opened'
      Visibility <- "20_TANKS_IP_DATA_RIO_01_FIRST_TANK_GTT_ISOL_VALVE_OPEN"
   Group "Group_1" at 120,420 size 35x38; Picture "Graphic_72"
   TextField "Text field_72" at 112,415 size 54x20; Text 'Closed'
      Visibility <- "20_TANKS_IP_DATA_RIO_07_FIRST_TANK_GTT_ISOL_VALVE_CLSD"
   TextField "Text field_73" at 112,415 size 54x20; Text 'Opened'
      Visibility <- "20_TANKS_IP_DATA_RIO_07_FIRST_TANK_GTT_ISOL_VALVE_OPEN"
   TextField "Text field_8" at 438,401 size 54x20; Text 'Closed'
      Visibility <- "20_TANKS_IP_DATA_RIO_05_FIRST_TANK_GTT_ISOL_VALVE_CLSD"
   TextField "Text field_9" at 438,401 size 54x20; Text 'Opened'
      Visibility <- "20_TANKS_IP_DATA_RIO_05_FIRST_TANK_GTT_ISOL_VALVE_OPEN"
   GraphicView "Graphic view_1" at 415,396 size 22x31; Picture "Graphic_162"
   TextField "Text field_10" at 438,482 size 54x20; Text 'Closed'
      Visibility <- "20_TANKS_IP_DATA_RIO_05_SECOND_TANK_GTT_ISOL_VALVE_CLSD"
   TextField "Text field_11" at 438,482 size 54x20; Text 'Opened'
      Visibility <- "20_TANKS_IP_DATA_RIO_05_SECOND_TANK_GTT_ISOL_VALVE_OPEN"
   GraphicView "Graphic view_3" at 415,476 size 22x31; Picture "Graphic_162"
   IOField "I/O field_5" at 441,560 size 72x20; FormatPattern 999; Unit Nm³/hr
      ProcessValue <- "20_TANKS_IP_DATA_RIO_05_SECOND_TANK_USD_FLOW"
   IOField "I/O field_6" at 441,599 size 72x20; FormatPattern 999; Unit Nm³/hr
      ProcessValue <- "20_TANKS_IP_DATA_RIO_05_SECOND_TANK_MBG_FLOW"
   TextField "Text field_12" at 395,602 size 29x14; Text 'MBG'
   TextField "Text field_13" at 417,545 size 33x15; Text 'USD'
   IOField "I/O field_7" at 441,289 size 72x20; FormatPattern 999; Unit Nm³/hr
      ProcessValue <- "20_TANKS_IP_DATA_RIO_05_FIRST_TANK_MBG_FLOW"
   IOField "I/O field_8" at 441,330 size 72x20; FormatPattern 999; Unit Nm³/hr
      ProcessValue <- "20_TANKS_IP_DATA_RIO_05_FIRST_TANK_USD_FLOW"
   TextField "Text field_14" at 393,291 size 34x14; Text 'MBG'
   TextField "Text field_15" at 416,349 size 28x14; Text 'USD'
   TextField "Text field_16" at 570,402 size 54x20; Text 'Closed'
      Visibility <- "20_TANKS_IP_DATA_RIO_04_FIRST_TANK_GTT_ISOL_VALVE_CLSD"
   TextField "Text field_17" at 570,402 size 54x20; Text 'Opened'
      Visibility <- "20_TANKS_IP_DATA_RIO_04_FIRST_TANK_GTT_ISOL_VALVE_OPEN"
   GraphicView "Graphic view_15" at 547,396 size 22x31; Picture "Graphic_162"
   TextField "Text field_18" at 570,482 size 54x20; Text 'Closed'
      Visibility <- "20_TANKS_IP_DATA_RIO_04_SECOND_TANK_GTT_ISOL_VALVE_CLSD"
   TextField "Text field_29" at 570,482 size 54x20; Text 'Opened'
      Visibility <- "20_TANKS_IP_DATA_RIO_04_SECOND_TANK_GTT_ISOL_VALVE_OPEN"
   GraphicView "Graphic view_16" at 547,476 size 22x31; Picture "Graphic_162"
   IOField "I/O field_9" at 573,560 size 72x20; FormatPattern 999; Unit Nm³/hr
      ProcessValue <- "20_TANKS_IP_DATA_RIO_04_SECOND_TANK_USD_FLOW"
   IOField "I/O field_10" at 573,599 size 72x20; FormatPattern 999; Unit Nm³/hr
      ProcessValue <- "20_TANKS_IP_DATA_RIO_04_SECOND_TANK_MBG_FLOW"
   TextField "Text field_30" at 527,602 size 29x14; Text 'MBG'
   TextField "Text field_31" at 549,545 size 33x15; Text 'USD'
   IOField "I/O field_11" at 573,289 size 72x20; FormatPattern 999; Unit Nm³/hr
      ProcessValue <- "20_TANKS_IP_DATA_RIO_04_FIRST_TANK_MBG_FLOW"
   IOField "I/O field_12" at 573,330 size 72x20; FormatPattern 999; Unit Nm³/hr
      ProcessValue <- "20_TANKS_IP_DATA_RIO_04_FIRST_TANK_USD_FLOW"
   TextField "Text field_32" at 525,291 size 34x14; Text 'MBG'
   TextField "Text field_33" at 548,349 size 28x14; Text 'USD'
   TextField "Text field_34" at 702,401 size 54x20; Text 'Closed'
      Visibility <- "20_TANKS_IP_DATA_RIO_03_FIRST_TANK_GTT_ISOL_VALVE_CLSD"
   TextField "Text field_35" at 702,401 size 54x20; Text 'Opened'
      Visibility <- "20_TANKS_IP_DATA_RIO_03_FIRST_TANK_GTT_ISOL_VALVE_OPEN"
   GraphicView "Graphic view_21" at 679,396 size 22x31; Picture "Graphic_162"
   TextField "Text field_36" at 702,482 size 54x20; Text 'Closed'
      Visibility <- "20_TANKS_IP_DATA_RIO_03_SECOND_TANK_GTT_ISOL_VALVE_CLSD"
   TextField "Text field_37" at 702,482 size 54x20; Text 'Opened'
      Visibility <- "20_TANKS_IP_DATA_RIO_03_SECOND_TANK_GTT_ISOL_VALVE_OPEN"
   GraphicView "Graphic view_22" at 679,476 size 22x31; Picture "Graphic_162"
   IOField "I/O field_13" at 705,560 size 72x20; FormatPattern 999; Unit Nm³/hr
      ProcessValue <- "20_TANKS_IP_DATA_RIO_03_SECOND_TANK_USD_FLOW"
   IOField "I/O field_14" at 705,599 size 72x20; FormatPattern 999; Unit Nm³/hr
      ProcessValue <- "20_TANKS_IP_DATA_RIO_03_SECOND_TANK_MBG_FLOW"
   TextField "Text field_38" at 659,602 size 29x14; Text 'MBG'
   TextField "Text field_39" at 681,545 size 33x15; Text 'USD'
   IOField "I/O field_15" at 705,289 size 72x20; FormatPattern 999; Unit Nm³/hr
      ProcessValue <- "20_TANKS_IP_DATA_RIO_03_FIRST_TANK_MBG_FLOW"
   IOField "I/O field_16" at 705,330 size 72x20; FormatPattern 999; Unit Nm³/hr
      ProcessValue <- "20_TANKS_IP_DATA_RIO_03_FIRST_TANK_USD_FLOW"
   TextField "Text field_40" at 657,291 size 34x14; Text 'MBG'
   TextField "Text field_41" at 680,349 size 28x14; Text 'USD'
   TextField "Text field_42" at 834,401 size 54x20; Text 'Closed'
      Visibility <- "20_TANKS_IP_DATA_RIO_02_FIRST_TANK_GTT_ISOL_VALVE_CLSD"
   TextField "Text field_43" at 834,401 size 54x20; Text 'Opened'
      Visibility <- "20_TANKS_IP_DATA_RIO_02_FIRST_TANK_GTT_ISOL_VALVE_OPEN"
   GraphicView "Graphic view_27" at 811,396 size 22x31; Picture "Graphic_162"
   TextField "Text field_44" at 834,482 size 54x20; Text 'Closed'
      Visibility <- "20_TANKS_IP_DATA_RIO_02_SECOND_TANK_GTT_ISOL_VALVE_CLSD"
   TextField "Text field_45" at 834,482 size 54x20; Text 'Opened'
      Visibility <- "20_TANKS_IP_DATA_RIO_02_SECOND_TANK_GTT_ISOL_VALVE_OPEN"
   GraphicView "Graphic view_28" at 811,476 size 22x31; Picture "Graphic_162"
   IOField "I/O field_17" at 837,560 size 72x20; FormatPattern 999; Unit Nm³/hr
      ProcessValue <- "20_TANKS_IP_DATA_RIO_02_SECOND_TANK_USD_FLOW"
   IOField "I/O field_18" at 837,599 size 72x20; FormatPattern 999; Unit Nm³/hr
      ProcessValue <- "20_TANKS_IP_DATA_RIO_02_SECOND_TANK_MBG_FLOW"
   TextField "Text field_46" at 791,602 size 29x14; Text 'MBG'
   TextField "Text field_47" at 813,545 size 33x15; Text 'USD'
   IOField "I/O field_19" at 837,289 size 72x20; FormatPattern 999; Unit Nm³/hr
      ProcessValue <- "20_TANKS_IP_DATA_RIO_02_FIRST_TANK_MBG_FLOW"
   IOField "I/O field_20" at 837,330 size 72x20; FormatPattern 999; Unit Nm³/hr
      ProcessValue <- "20_TANKS_IP_DATA_RIO_02_FIRST_TANK_USD_FLOW"
   TextField "Text field_48" at 789,291 size 34x14; Text 'MBG'
   TextField "Text field_49" at 812,349 size 28x14; Text 'USD'
   TextField "Text field_50" at 966,401 size 54x20; Text 'Closed'
      Visibility <- "20_TANKS_IP_DATA_RIO_01_SECOND_TANK_GTT_ISOL_VALVE_CLSD"
   TextField "Text field_51" at 966,401 size 54x20; Text 'Opened'
      Visibility <- "20_TANKS_IP_DATA_RIO_01_SECOND_TANK_GTT_ISOL_VALVE_OPEN"
   GraphicView "Graphic view_33" at 943,396 size 22x31; Picture "Graphic_162"
   TextField "Text field_52" at 966,482 size 54x20; Text 'Closed'
      Visibility <- "20_TANKS_IP_DATA_RIO_01_THIRD_TANK_GTT_ISOL_VALVE_CLSD"
   TextField "Text field_53" at 966,482 size 54x20; Text 'Opened'
      Visibility <- "20_TANKS_IP_DATA_RIO_01_THIRD_TANK_GTT_ISOL_VALVE_OPEN"
   GraphicView "Graphic view_34" at 943,476 size 22x31; Picture "Graphic_162"
   IOField "I/O field_21" at 969,560 size 72x20; FormatPattern 999; Unit Nm³/hr
      ProcessValue <- "20_TANKS_IP_DATA_RIO_01_THIRD_TANK_USD_FLOW"
   IOField "I/O field_22" at 969,599 size 72x20; FormatPattern 999; Unit Nm³/hr
      ProcessValue <- "20_TANKS_IP_DATA_RIO_01_THIRD_TANK_MBG_FLOW"
   TextField "Text field_54" at 923,602 size 29x14; Text 'MBG'
   TextField "Text field_55" at 945,545 size 33x15; Text 'USD'
   IOField "I/O field_23" at 969,289 size 72x20; FormatPattern 999; Unit Nm³/hr
      ProcessValue <- "20_TANKS_IP_DATA_RIO_01_SECOND_TANK_MBG_FLOW"
   IOField "I/O field_24" at 969,330 size 72x20; FormatPattern 999; Unit Nm³/hr
      ProcessValue <- "20_TANKS_IP_DATA_RIO_01_SECOND_TANK_USD_FLOW"
   TextField "Text field_56" at 921,291 size 34x14; Text 'MBG'
   TextField "Text field_57" at 944,349 size 28x14; Text 'USD'
   GraphicView "Graphic view_17" at 575,446 size 485x12; Picture "Graphic_151"
   Button "Button_13" at 252,437 size 37x30; TextOff 'DB&B'
   TextField "Text field_58" at 188,226 size 50x40; Text 'Safe Area'
   TextField "Text field_59" at 417,454 size 137x22; Text 'Hazardous Area'
   Button "HmiScreenItemData_5" at 180,144 size 116x50; TextOn 'Back'; TextOff 'Tank Status'
      on Release: function_efd93a16("Tank Status", 400, 250, -1, -1, 1)
   IOField "I/O field_25" at 100,385 size 72x20; FormatPattern 999; Unit Nm³/hr
      ProcessValue <- "20_TANKS_IP_DATA_RIO_07_FIRST_TANK_MBG_FLOW"
   IOField "I/O field_26" at 100,491 size 72x20; FormatPattern 999; Unit Nm³/hr
      ProcessValue <- "20_TANKS_IP_DATA_RIO_07_FIRST_TANK_USD_FLOW"
   TextField "Text field_66" at 107,527 size 34x14; Text 'USD'
   TextField "Text field_67" at 107,356 size 34x14; Text 'MBG'
   IOField "I/O field_27" at 1080,381 size 72x20; FormatPattern 999; Unit Nm³/hr
      ProcessValue <- "20_TANKS_IP_DATA_RIO_01_FIRST_TANK_MBG_FLOW"
   IOField "I/O field_28" at 1080,491 size 72x20; FormatPattern 999; Unit Nm³/hr
      ProcessValue <- "20_TANKS_IP_DATA_RIO_01_FIRST_TANK_USD_FLOW"
   TextField "Text field_68" at 1111,527 size 34x14; Text 'USD'
   TextField "Text field_69" at 1111,350 size 34x14; Text 'MBG'
   Button "Button_20" at 724,152 size 115x34; TextOff 'Re-Oxygenation'
      Appearance <- "2110_BTCS_CNTRL_DB_BTCS_STEP"
   Button "Button_21" at 845,152 size 93x34; TextOff 'Post Dwell'
      Appearance <- "2110_BTCS_CNTRL_DB_BTCS_STATE"
   Circle "Circle_1" at 137,105 size 29x29
      Appearance <- "2110_BTCS_CNTRL_DB_BTCS_STATE"
   Circle "Circle_8" at 775,89 size 14x14
      Appearance <- "100_GCU_AUTO_SEQ_DB_CRNT_STEP"
   Circle "Circle_9" at 685,89 size 14x14
      Appearance <- "100_GCU_AUTO_SEQ_DB_CRNT_STEP"
   Circle "Circle_11" at 595,89 size 14x14
      Appearance <- "51_SLAVE_STATUS_RUNNING"